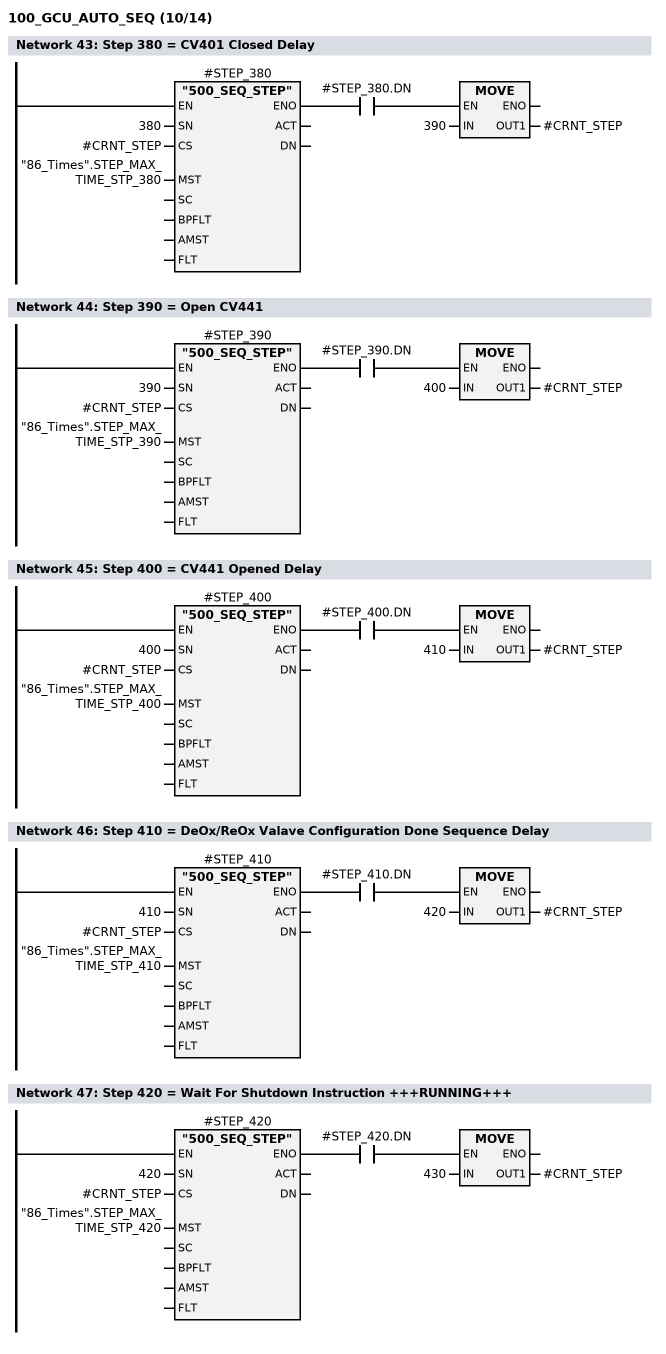
   RUNG wire#powerrail
      #STEP_380(SN := 380, CS := #CRNT_STEP, MST := "86_Times".STEP_MAX_TIME_STP_380, SC :=, BPFLT :=, AMST :=, FLT :=, ACT =>, DN =>)
      Contact( #STEP_380.DN )
      Move(in := 390, out1 => #CRNT_STEP)
   END_RUNG
   // the same network as SCL:
   #STEP_380(SN := 380, CS := #CRNT_STEP, MST := "86_Times".STEP_MAX_TIME_STP_380, ENO => #_w1);   // "500_SEQ_STEP"
   IF #_w1 AND #STEP_380.DN THEN #CRNT_STEP := 390; END_IF;
END_REGION

REGION Network 44: Step 390 = Open CV441
   RUNG wire#powerrail
      #STEP_390(SN := 390, CS := #CRNT_STEP, MST := "86_Times".STEP_MAX_TIME_STP_390, SC :=, BPFLT :=, AMST :=, FLT :=, ACT =>, DN =>)
      Contact( #STEP_390.DN )
      Move(in := 400, out1 => #CRNT_STEP)
   END_RUNG
   // the same network as SCL:
   #STEP_390(SN := 390, CS := #CRNT_STEP, MST := "86_Times".STEP_MAX_TIME_STP_390, ENO => #_w1);   // "500_SEQ_STEP"
   IF #_w1 AND #STEP_390.DN THEN #CRNT_STEP := 400; END_IF;
END_REGION

REGION Network 45: Step 400 = CV441 Opened Delay
   RUNG wire#powerrail
      #STEP_400(SN := 400, CS := #CRNT_STEP, MST := "86_Times".STEP_MAX_TIME_STP_400, SC :=, BPFLT :=, AMST :=, FLT :=, ACT =>, DN =>)
      Contact( #STEP_400.DN )
      Move(in := 410, out1 => #CRNT_STEP)
   END_RUNG
   // the same network as SCL:
   #STEP_400(SN := 400, CS := #CRNT_STEP, MST := "86_Times".STEP_MAX_TIME_STP_400, ENO => #_w1);   // "500_SEQ_STEP"
   IF #_w1 AND #STEP_400.DN THEN #CRNT_STEP := 410; END_IF;
END_REGION

REGION Network 46: Step 410 = DeOx/ReOx Valave Configuration Done Sequence Delay
   RUNG wire#powerrail
      #STEP_410(SN := 410, CS := #CRNT_STEP, MST := "86_Times".STEP_MAX_TIME_STP_410, SC :=, BPFLT :=, AMST :=, FLT :=, ACT =>, DN =>)
      Contact( #STEP_410.DN )
      Move(in := 420, out1 => #CRNT_STEP)
   END_RUNG
   // the same network as SCL:
   #STEP_410(SN := 410, CS := #CRNT_STEP, MST := "86_Times".STEP_MAX_TIME_STP_410, ENO => #_w1);   // "500_SEQ_STEP"
   IF #_w1 AND #STEP_410.DN THEN #CRNT_STEP := 420; END_IF;
END_REGION

REGION Network 47: Step 420 = Wait For Shutdown Instruction +++RUNNING+++
   RUNG wire#powerrail
      #STEP_420(SN := 420, CS := #CRNT_STEP, MST := "86_Times".STEP_MAX_TIME_STP_420, SC :=, BPFLT :=, AMST :=, FLT :=, ACT =>, DN =>)
      Contact( #STEP_420.DN )
      Move(in := 430, out1 => #CRNT_STEP)
   END_RUNG
   // the same network as SCL:
   #STEP_420(SN := 420, CS := #CRNT_STEP, MST := "86_Times".STEP_MAX_TIME_STP_420, ENO => #_w1);   // "500_SEQ_STEP"
   IF #_w1 AND #STEP_420.DN THEN #CRNT_STEP := 430; END_IF;
END_REGION

REGION Network 48: Step 430 = Spare Step (Not Used)
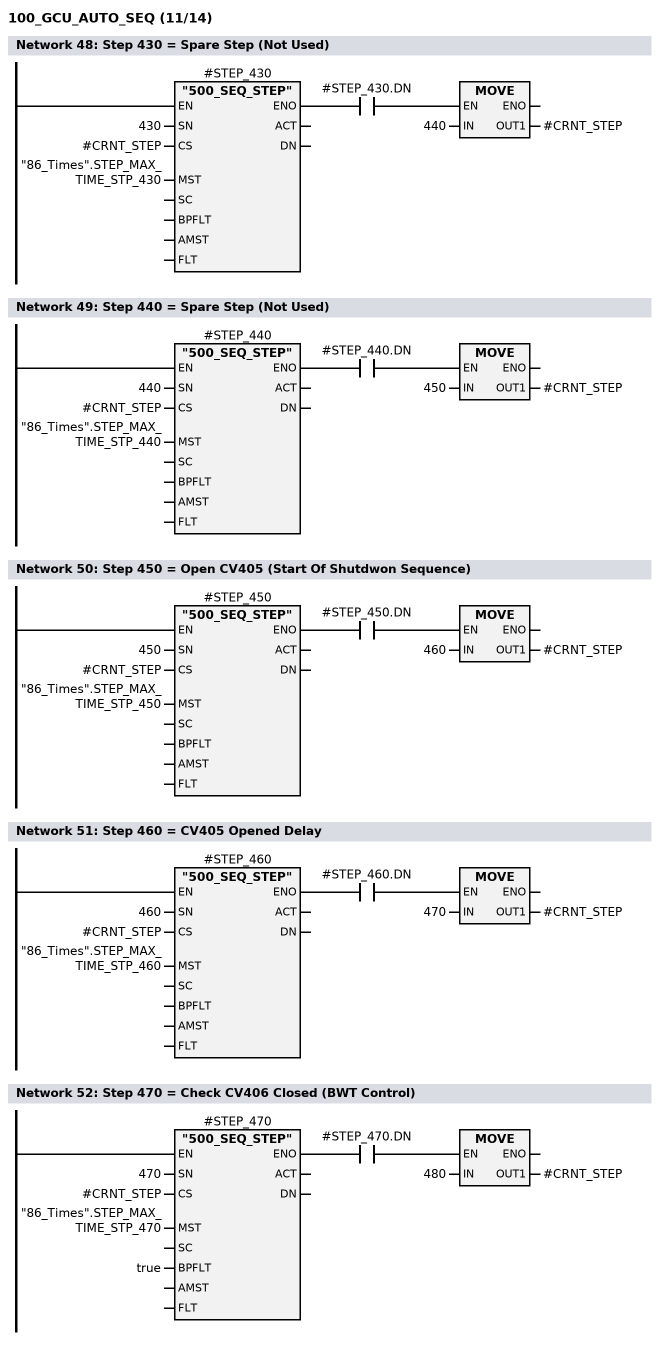
   RUNG wire#powerrail
      #STEP_430(SN := 430, CS := #CRNT_STEP, MST := "86_Times".STEP_MAX_TIME_STP_430, SC :=, BPFLT :=, AMST :=, FLT :=, ACT =>, DN =>)
      Contact( #STEP_430.DN )
      Move(in := 440, out1 => #CRNT_STEP)
   END_RUNG
   // the same network as SCL:
   #STEP_430(SN := 430, CS := #CRNT_STEP, MST := "86_Times".STEP_MAX_TIME_STP_430, ENO => #_w1);   // "500_SEQ_STEP"
   IF #_w1 AND #STEP_430.DN THEN #CRNT_STEP := 440; END_IF;
END_REGION

REGION Network 49: Step 440 = Spare Step (Not Used)
   RUNG wire#powerrail
      #STEP_440(SN := 440, CS := #CRNT_STEP, MST := "86_Times".STEP_MAX_TIME_STP_440, SC :=, BPFLT :=, AMST :=, FLT :=, ACT =>, DN =>)
      Contact( #STEP_440.DN )
      Move(in := 450, out1 => #CRNT_STEP)
   END_RUNG
   // the same network as SCL:
   #STEP_440(SN := 440, CS := #CRNT_STEP, MST := "86_Times".STEP_MAX_TIME_STP_440, ENO => #_w1);   // "500_SEQ_STEP"
   IF #_w1 AND #STEP_440.DN THEN #CRNT_STEP := 450; END_IF;
END_REGION

REGION Network 50: Step 450 = Open CV405 (Start Of Shutdwon Sequence)
   RUNG wire#powerrail
      #STEP_450(SN := 450, CS := #CRNT_STEP, MST := "86_Times".STEP_MAX_TIME_STP_450, SC :=, BPFLT :=, AMST :=, FLT :=, ACT =>, DN =>)
      Contact( #STEP_450.DN )
      Move(in := 460, out1 => #CRNT_STEP)
   END_RUNG
   // the same network as SCL:
   #STEP_450(SN := 450, CS := #CRNT_STEP, MST := "86_Times".STEP_MAX_TIME_STP_450, ENO => #_w1);   // "500_SEQ_STEP"
   IF #_w1 AND #STEP_450.DN THEN #CRNT_STEP := 460; END_IF;
END_REGION

REGION Network 51: Step 460 = CV405 Opened Delay
   RUNG wire#powerrail
      #STEP_460(SN := 460, CS := #CRNT_STEP, MST := "86_Times".STEP_MAX_TIME_STP_460, SC :=, BPFLT :=, AMST :=, FLT :=, ACT =>, DN =>)
      Contact( #STEP_460.DN )
      Move(in := 470, out1 => #CRNT_STEP)
   END_RUNG
   // the same network as SCL:
   #STEP_460(SN := 460, CS := #CRNT_STEP, MST := "86_Times".STEP_MAX_TIME_STP_460, ENO => #_w1);   // "500_SEQ_STEP"
   IF #_w1 AND #STEP_460.DN THEN #CRNT_STEP := 470; END_IF;
END_REGION

REGION Network 52: Step 470 = Check CV406 Closed (BWT Control)
   RUNG wire#powerrail
      #STEP_470(SN := 470, CS := #CRNT_STEP, MST := "86_Times".STEP_MAX_TIME_STP_470, SC :=, BPFLT := true, AMST :=, FLT :=, ACT =>, DN =>)
      Contact( #STEP_470.DN )
      Move(in := 480, out1 => #CRNT_STEP)
   END_RUNG
   // the same network as SCL:
   #STEP_470(SN := 470, CS := #CRNT_STEP, MST := "86_Times".STEP_MAX_TIME_STP_470, BPFLT := true, ENO => #_w1);   // "500_SEQ_STEP"
   IF #_w1 AND #STEP_470.DN THEN #CRNT_STEP := 480; END_IF;
END_REGION

REGION Network 53: Step 480 = CV406 Closed Delay
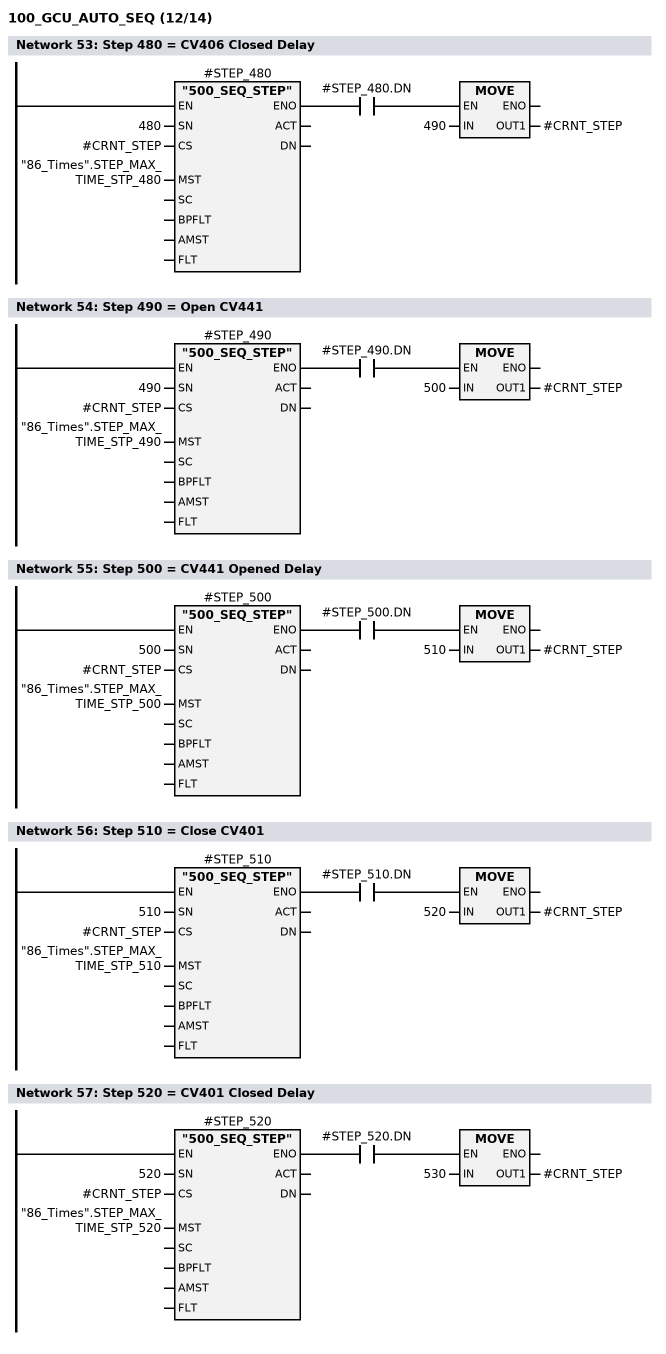
   RUNG wire#powerrail
      #STEP_480(SN := 480, CS := #CRNT_STEP, MST := "86_Times".STEP_MAX_TIME_STP_480, SC :=, BPFLT :=, AMST :=, FLT :=, ACT =>, DN =>)
      Contact( #STEP_480.DN )
      Move(in := 490, out1 => #CRNT_STEP)
   END_RUNG
   // the same network as SCL:
   #STEP_480(SN := 480, CS := #CRNT_STEP, MST := "86_Times".STEP_MAX_TIME_STP_480, ENO => #_w1);   // "500_SEQ_STEP"
   IF #_w1 AND #STEP_480.DN THEN #CRNT_STEP := 490; END_IF;
END_REGION

REGION Network 54: Step 490 = Open CV441
   RUNG wire#powerrail
      #STEP_490(SN := 490, CS := #CRNT_STEP, MST := "86_Times".STEP_MAX_TIME_STP_490, SC :=, BPFLT :=, AMST :=, FLT :=, ACT =>, DN =>)
      Contact( #STEP_490.DN )
      Move(in := 500, out1 => #CRNT_STEP)
   END_RUNG
   // the same network as SCL:
   #STEP_490(SN := 490, CS := #CRNT_STEP, MST := "86_Times".STEP_MAX_TIME_STP_490, ENO => #_w1);   // "500_SEQ_STEP"
   IF #_w1 AND #STEP_490.DN THEN #CRNT_STEP := 500; END_IF;
END_REGION

REGION Network 55: Step 500 = CV441 Opened Delay
   RUNG wire#powerrail
      #STEP_500(SN := 500, CS := #CRNT_STEP, MST := "86_Times".STEP_MAX_TIME_STP_500, SC :=, BPFLT :=, AMST :=, FLT :=, ACT =>, DN =>)
      Contact( #STEP_500.DN )
      Move(in := 510, out1 => #CRNT_STEP)
   END_RUNG
   // the same network as SCL:
   #STEP_500(SN := 500, CS := #CRNT_STEP, MST := "86_Times".STEP_MAX_TIME_STP_500, ENO => #_w1);   // "500_SEQ_STEP"
   IF #_w1 AND #STEP_500.DN THEN #CRNT_STEP := 510; END_IF;
END_REGION

REGION Network 56: Step 510 = Close CV401
   RUNG wire#powerrail
      #STEP_510(SN := 510, CS := #CRNT_STEP, MST := "86_Times".STEP_MAX_TIME_STP_510, SC :=, BPFLT :=, AMST :=, FLT :=, ACT =>, DN =>)
      Contact( #STEP_510.DN )
      Move(in := 520, out1 => #CRNT_STEP)
   END_RUNG
   // the same network as SCL:
   #STEP_510(SN := 510, CS := #CRNT_STEP, MST := "86_Times".STEP_MAX_TIME_STP_510, ENO => #_w1);   // "500_SEQ_STEP"
   IF #_w1 AND #STEP_510.DN THEN #CRNT_STEP := 520; END_IF;
END_REGION

REGION Network 57: Step 520 = CV401 Closed Delay
   RUNG wire#powerrail
      #STEP_520(SN := 520, CS := #CRNT_STEP, MST := "86_Times".STEP_MAX_TIME_STP_520, SC :=, BPFLT :=, AMST :=, FLT :=, ACT =>, DN =>)
      Contact( #STEP_520.DN )
      Move(in := 530, out1 => #CRNT_STEP)
   END_RUNG
   // the same network as SCL:
   #STEP_520(SN := 520, CS := #CRNT_STEP, MST := "86_Times".STEP_MAX_TIME_STP_520, ENO => #_w1);   // "500_SEQ_STEP"
   IF #_w1 AND #STEP_520.DN THEN #CRNT_STEP := 530; END_IF;
END_REGION

REGION Network 58: Step 530 = Stop E400
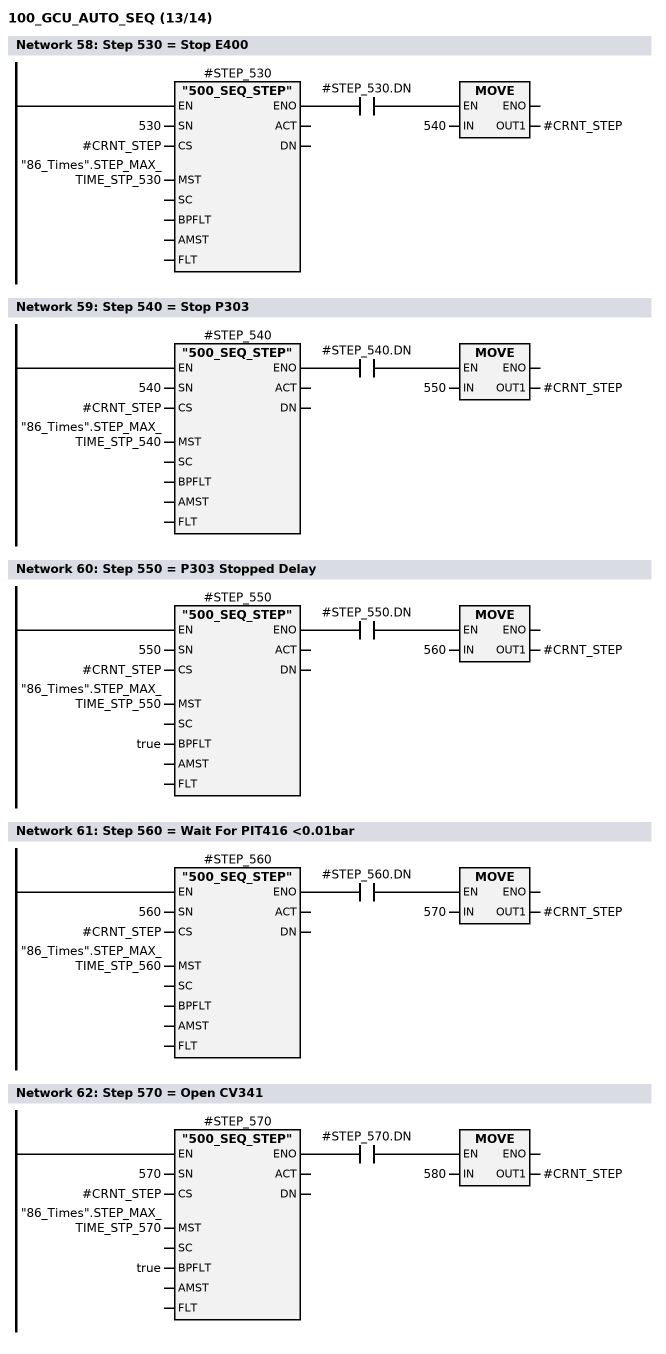
   RUNG wire#powerrail
      #STEP_530(SN := 530, CS := #CRNT_STEP, MST := "86_Times".STEP_MAX_TIME_STP_530, SC :=, BPFLT :=, AMST :=, FLT :=, ACT =>, DN =>)
      Contact( #STEP_530.DN )
      Move(in := 540, out1 => #CRNT_STEP)
   END_RUNG
   // the same network as SCL:
   #STEP_530(SN := 530, CS := #CRNT_STEP, MST := "86_Times".STEP_MAX_TIME_STP_530, ENO => #_w1);   // "500_SEQ_STEP"
   IF #_w1 AND #STEP_530.DN THEN #CRNT_STEP := 540; END_IF;
END_REGION

REGION Network 59: Step 540 = Stop P303
   RUNG wire#powerrail
      #STEP_540(SN := 540, CS := #CRNT_STEP, MST := "86_Times".STEP_MAX_TIME_STP_540, SC :=, BPFLT :=, AMST :=, FLT :=, ACT =>, DN =>)
      Contact( #STEP_540.DN )
      Move(in := 550, out1 => #CRNT_STEP)
   END_RUNG
   // the same network as SCL:
   #STEP_540(SN := 540, CS := #CRNT_STEP, MST := "86_Times".STEP_MAX_TIME_STP_540, ENO => #_w1);   // "500_SEQ_STEP"
   IF #_w1 AND #STEP_540.DN THEN #CRNT_STEP := 550; END_IF;
END_REGION

REGION Network 60: Step 550 = P303 Stopped Delay
   RUNG wire#powerrail
      #STEP_550(SN := 550, CS := #CRNT_STEP, MST := "86_Times".STEP_MAX_TIME_STP_550, SC :=, BPFLT := true, AMST :=, FLT :=, ACT =>, DN =>)
      Contact( #STEP_550.DN )
      Move(in := 560, out1 => #CRNT_STEP)
   END_RUNG
   // the same network as SCL:
   #STEP_550(SN := 550, CS := #CRNT_STEP, MST := "86_Times".STEP_MAX_TIME_STP_550, BPFLT := true, ENO => #_w1);   // "500_SEQ_STEP"
   IF #_w1 AND #STEP_550.DN THEN #CRNT_STEP := 560; END_IF;
END_REGION

REGION Network 61: Step 560 = Wait For PIT416 <0.01bar
   RUNG wire#powerrail
      #STEP_560(SN := 560, CS := #CRNT_STEP, MST := "86_Times".STEP_MAX_TIME_STP_560, SC :=, BPFLT :=, AMST :=, FLT :=, ACT =>, DN =>)
      Contact( #STEP_560.DN )
      Move(in := 570, out1 => #CRNT_STEP)
   END_RUNG
   // the same network as SCL:
   #STEP_560(SN := 560, CS := #CRNT_STEP, MST := "86_Times".STEP_MAX_TIME_STP_560, ENO => #_w1);   // "500_SEQ_STEP"
   IF #_w1 AND #STEP_560.DN THEN #CRNT_STEP := 570; END_IF;
END_REGION

REGION Network 62: Step 570 = Open CV341
   RUNG wire#powerrail
      #STEP_570(SN := 570, CS := #CRNT_STEP, MST := "86_Times".STEP_MAX_TIME_STP_570, SC :=, BPFLT := true, AMST :=, FLT :=, ACT =>, DN =>)
      Contact( #STEP_570.DN )
      Move(in := 580, out1 => #CRNT_STEP)
   END_RUNG
   // the same network as SCL:
   #STEP_570(SN := 570, CS := #CRNT_STEP, MST := "86_Times".STEP_MAX_TIME_STP_570, BPFLT := true, ENO => #_w1);   // "500_SEQ_STEP"
   IF #_w1 AND #STEP_570.DN THEN #CRNT_STEP := 580; END_IF;
END_REGION

REGION Network 63: Step 580 = CV341 Opened Delay
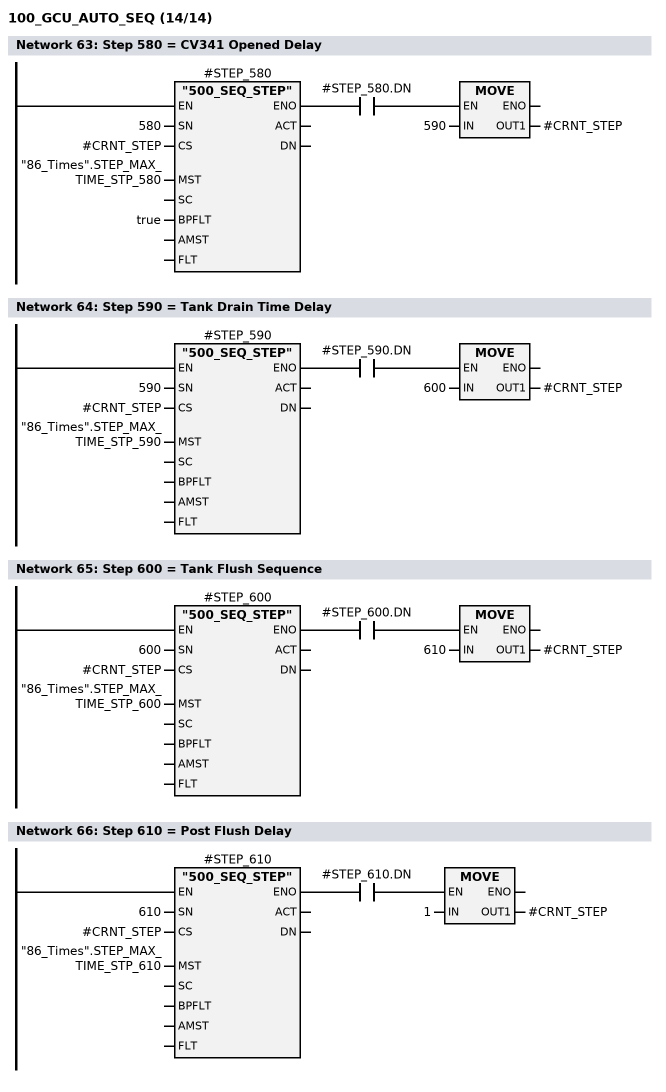
   RUNG wire#powerrail
      #STEP_580(SN := 580, CS := #CRNT_STEP, MST := "86_Times".STEP_MAX_TIME_STP_580, SC :=, BPFLT := true, AMST :=, FLT :=, ACT =>, DN =>)
      Contact( #STEP_580.DN )
      Move(in := 590, out1 => #CRNT_STEP)
   END_RUNG
   // the same network as SCL:
   #STEP_580(SN := 580, CS := #CRNT_STEP, MST := "86_Times".STEP_MAX_TIME_STP_580, BPFLT := true, ENO => #_w1);   // "500_SEQ_STEP"
   IF #_w1 AND #STEP_580.DN THEN #CRNT_STEP := 590; END_IF;
END_REGION

REGION Network 64: Step 590 = Tank Drain Time Delay
   RUNG wire#powerrail
      #STEP_590(SN := 590, CS := #CRNT_STEP, MST := "86_Times".STEP_MAX_TIME_STP_590, SC :=, BPFLT :=, AMST :=, FLT :=, ACT =>, DN =>)
      Contact( #STEP_590.DN )
      Move(in := 600, out1 => #CRNT_STEP)
   END_RUNG
   // the same network as SCL:
   #STEP_590(SN := 590, CS := #CRNT_STEP, MST := "86_Times".STEP_MAX_TIME_STP_590, ENO => #_w1);   // "500_SEQ_STEP"
   IF #_w1 AND #STEP_590.DN THEN #CRNT_STEP := 600; END_IF;
END_REGION

REGION Network 65: Step 600 = Tank Flush Sequence
   RUNG wire#powerrail
      #STEP_600(SN := 600, CS := #CRNT_STEP, MST := "86_Times".STEP_MAX_TIME_STP_600, SC :=, BPFLT :=, AMST :=, FLT :=, ACT =>, DN =>)
      Contact( #STEP_600.DN )
      Move(in := 610, out1 => #CRNT_STEP)
   END_RUNG
   // the same network as SCL:
   #STEP_600(SN := 600, CS := #CRNT_STEP, MST := "86_Times".STEP_MAX_TIME_STP_600, ENO => #_w1);   // "500_SEQ_STEP"
   IF #_w1 AND #STEP_600.DN THEN #CRNT_STEP := 610; END_IF;
END_REGION

REGION Network 66: Step 610 = Post Flush Delay
   RUNG wire#powerrail
      #STEP_610(SN := 610, CS := #CRNT_STEP, MST := "86_Times".STEP_MAX_TIME_STP_610, SC :=, BPFLT :=, AMST :=, FLT :=, ACT =>, DN =>)
      Contact( #STEP_610.DN )
      Move(in := 1, out1 => #CRNT_STEP)
   END_RUNG
   // the same network as SCL:
   #STEP_610(SN := 610, CS := #CRNT_STEP, MST := "86_Times".STEP_MAX_TIME_STP_610, ENO => #_w1);   // "500_SEQ_STEP"
   IF #_w1 AND #STEP_610.DN THEN #CRNT_STEP := 1; END_IF;
END_REGION
END_FUNCTION_BLOCK

FUNCTION_BLOCK "Setpoint Override"   // FB104, LAD
{ S7_Optimized_Access := 'TRUE' }
VERSION : 0.1
   VAR_INPUT
      Enable : Bool;
      "Activate Temp Prot" : Bool := true;
      Temperature : Real;
      "Temperature Setpoint" : Real := 250.0;
      "Temperature Tolerance" : Real := 10.0;
      "Activate Press Prot" : Bool;
      Pressure : Real;
      "Pressure Setpoint" : Real := 5.0;
      "Pressure Tolerance" : Real := 0.2;
      "Pressure Target" : Real := 3.5;
      "Pressure Safe Target" : Real := 3.0;
      "Activate Tank Change Prot" : Bool := true;
      "Tank Change TimeOut" : Time := T#60s;
      "Tank Change" : Bool := true;
      Reset : Bool;
   END_VAR
   VAR_OUTPUT
      "Pressure Target Override" : Real;
      "Pressure Safe Override" : Real;
   END_VAR
   VAR
      "Temperature Setpoint Aux" : Real;
      "Pressure Setpoint Aux" : Real;
      "Set Pressure" : Bool;
      "Set Pressure Aux" : Bool;
      "Set Pressure by Temp" : Bool;
      "Set Pressure by Press" : Bool;
      "Set Pressure by Tank" : Bool;
   END_VAR
   VAR RETAIN
      "Pressure Target Memory" : Real;
   END_VAR
   VAR
      "Set Pressure Puls1" : Bool;
      "Set Pressure Puls2" : Bool;
      "Tank Change Protection" : TOF_TIME;
      "Pressure Protection" : TOF_TIME;
      "Pressure Memory Recover" : TON_TIME;
   END_VAR
   VAR_TEMP   // added for the SCL form of the ladder/FBD networks
      _w1 : Bool;
   END_VAR
BEGIN

REGION Network 1: Pressure Safe Corection
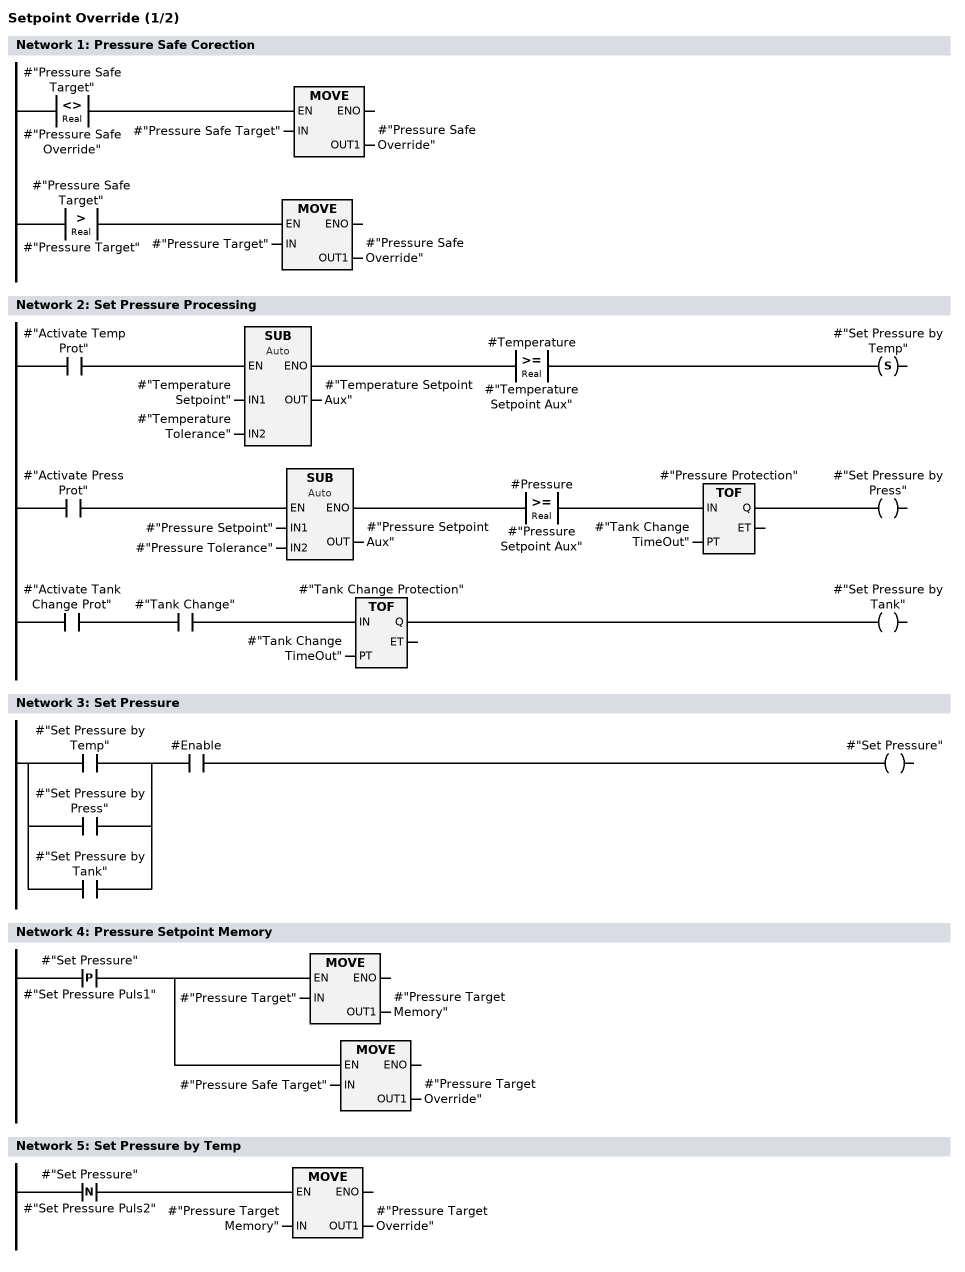
   RUNG wire#powerrail
      { S7_Templates := "SrcType := Real" } NE_Contact(in1 := #"Pressure Safe Target", in2 := #"Pressure Safe Override")
      Move(in := #"Pressure Safe Target", out1 => #"Pressure Safe Override")
   END_RUNG
   RUNG wire#powerrail
      { S7_Templates := "SrcType := Real" } GT_Contact(in1 := #"Pressure Safe Target", in2 := #"Pressure Target")
      Move(in := #"Pressure Target", out1 => #"Pressure Safe Override")
   END_RUNG
   // the same network as SCL:
   IF #"Pressure Safe Target" <> #"Pressure Safe Override" THEN
       #"Pressure Safe Override" := #"Pressure Safe Target";
   END_IF;
   IF #"Pressure Safe Target" > #"Pressure Target" THEN
       #"Pressure Safe Override" := #"Pressure Target";
   END_IF;
END_REGION

REGION Network 2: Set Pressure Processing
   IF #"Activate Temp Prot" THEN
       #"Temperature Setpoint Aux" := #"Temperature Setpoint" - #"Temperature Tolerance";
   END_IF;
   IF #"Activate Temp Prot" AND (#Temperature >= #"Temperature Setpoint Aux") THEN
       #"Set Pressure by Temp" := TRUE;
   END_IF;
   IF #"Activate Press Prot" THEN
       #"Pressure Setpoint Aux" := #"Pressure Setpoint" - #"Pressure Tolerance";
   END_IF;
   #"Pressure Protection"(IN := #"Activate Press Prot" AND (#Pressure >= #"Pressure Setpoint Aux"),   // TOF
                          PT := #"Tank Change TimeOut");
   #"Set Pressure by Press" := #"Pressure Protection".Q;
   #"Tank Change Protection"(IN := #"Activate Tank Change Prot" AND #"Tank Change",   // TOF
                           PT := #"Tank Change TimeOut");
   #"Set Pressure by Tank" := #"Tank Change Protection".Q;
END_REGION

REGION Network 3: Set Pressure
   RUNG wire#powerrail
      Contact( #"Set Pressure by Temp" )
      wire#w1
      Contact( #Enable )
      Coil( #"Set Pressure" )
   END_RUNG
   RUNG wire#powerrail
      Contact( #"Set Pressure by Press" )
   END_RUNG wire#w1
   RUNG wire#powerrail
      Contact( #"Set Pressure by Tank" )
   END_RUNG wire#w1
   // the same network as SCL:
   #"Set Pressure" := (#"Set Pressure by Temp" OR #"Set Pressure by Press" OR #"Set Pressure by Tank") AND #Enable;
END_REGION

REGION Network 4: Pressure Setpoint Memory
   RUNG wire#powerrail
      P_Contact(operand := #"Set Pressure", bit := #"Set Pressure Puls1")
      wire#w1
      Move(in := #"Pressure Target", out1 => #"Pressure Target Memory")
   END_RUNG
   RUNG wire#w1
      Move(in := #"Pressure Safe Target", out1 => #"Pressure Target Override")
   END_RUNG
   // the same network as SCL:
   #_w1 := #"Set Pressure" AND NOT #"Set Pressure Puls1";   // rising edge of #"Set Pressure"
   #"Set Pressure Puls1" := #"Set Pressure";
   IF #_w1 THEN
       #"Pressure Target Memory" := #"Pressure Target";
       #"Pressure Target Override" := #"Pressure Safe Target";
   END_IF;
END_REGION

REGION Network 5: Set Pressure by Temp
   RUNG wire#powerrail
      N_Contact(operand := #"Set Pressure", bit := #"Set Pressure Puls2")
      Move(in := #"Pressure Target Memory", out1 => #"Pressure Target Override")
   END_RUNG
   // the same network as SCL:
   #_w1 := NOT #"Set Pressure" AND #"Set Pressure Puls2";   // falling edge of #"Set Pressure"
   #"Set Pressure Puls2" := #"Set Pressure";
   IF #_w1 THEN #"Pressure Target Override" := #"Pressure Target Memory"; END_IF;
END_REGION

REGION Network 6: Set Pressure Back
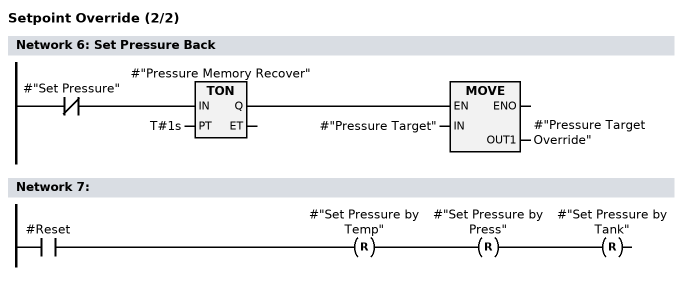
   #"Pressure Memory Recover"(IN := NOT #"Set Pressure", PT := T#1s);   // TON
   IF #"Pressure Memory Recover".Q THEN #"Pressure Target Override" := #"Pressure Target"; END_IF;
END_REGION

REGION Network 7
   RUNG wire#powerrail
      Contact( #Reset )
      R_Coil( #"Set Pressure by Temp" )
      R_Coil( #"Set Pressure by Press" )
      R_Coil( #"Set Pressure by Tank" )
   END_RUNG
   // the same network as SCL:
   IF #Reset THEN
       #"Set Pressure by Temp" := FALSE;
       #"Set Pressure by Press" := FALSE;
       #"Set Pressure by Tank" := FALSE;
   END_IF;
END_REGION
END_FUNCTION_BLOCK

FUNCTION_BLOCK "108_GCU_TNK_REFILL_SEQ"   // FB108, LAD
TITLE = GCU Tank Refill Sequence
{ S7_Optimized_Access := 'TRUE' }
AUTHOR : JRS
VERSION : 0.1
// For the automatic refilling of the GCU tank to the required level
   VAR_INPUT
      RUN : Bool;   // Block control
      LEVEL : Real;   // Tank level value
      TARGET : Real;   // Target level value
      LOW : Real;   // Low level value
      P305_PRSNT : Bool;   // P305 Fitted
      P305_RNG : Bool;   // Pump running
      P304_RNG : Bool;   // Pump running
      CV358_OPN : Bool;   // Valve open
      CV358_CLSD : Bool;   // Valve closed
   END_VAR
   VAR_OUTPUT
      RUN_P305 : Bool;   // Pump control
      RUN_P304 : Bool;   // Pump control
      OPEN_CV358 : Bool;   // Valve control
      FILLING : Bool;   // Filling status
   END_VAR
   VAR
      INTO_RUN_PLS : Bool;   // Pulse bit
      "STEP" : Int;   // Step number
      RNG : Bool;   // Running bit
      OUT_RUN_PLS : Bool;   // Pulse bit
   END_VAR
   VAR_TEMP   // added for the SCL form of the ladder/FBD networks
      _w1 : Bool;
   END_VAR
BEGIN

REGION Network 1: First Into Run
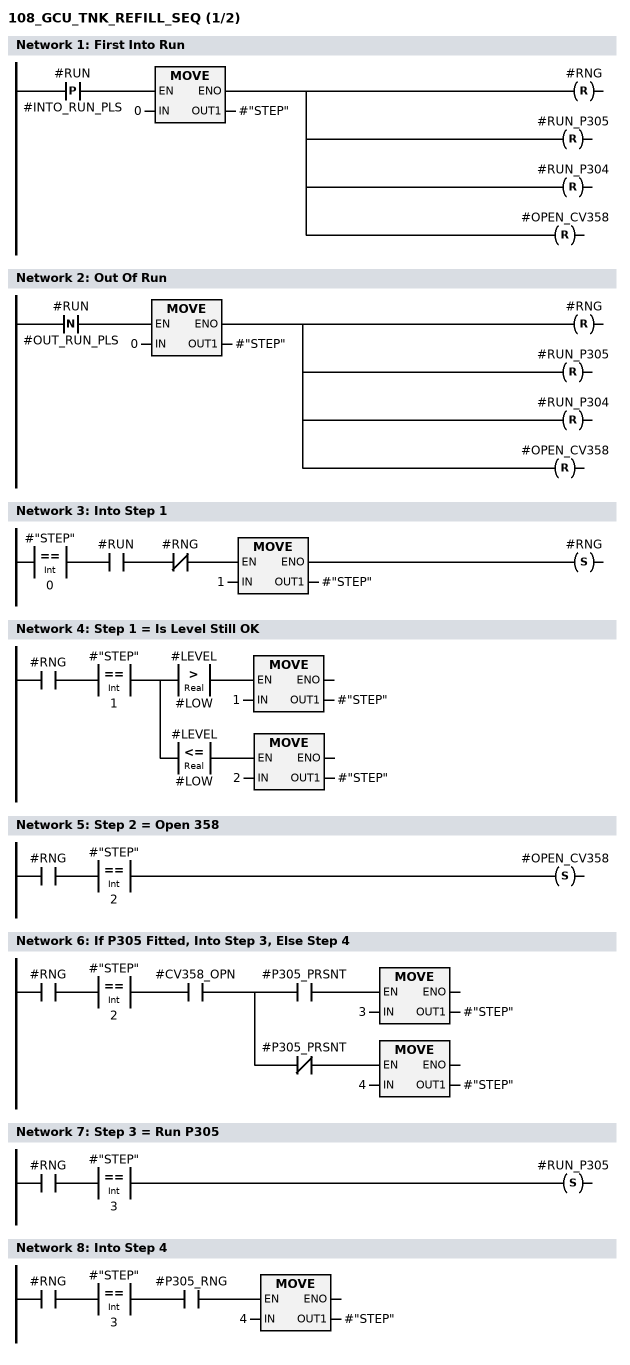
   RUNG wire#powerrail
      P_Contact(operand := #RUN, bit := #INTO_RUN_PLS)
      Move(in := 0, out1 => #"STEP")
      wire#w1
      R_Coil( #RNG )
   END_RUNG
   RUNG wire#w1
      R_Coil( #RUN_P305 )
   END_RUNG
   RUNG wire#w1
      R_Coil( #RUN_P304 )
   END_RUNG
   RUNG wire#w1
      R_Coil( #OPEN_CV358 )
   END_RUNG
   // the same network as SCL:
   #_w1 := #RUN AND NOT #INTO_RUN_PLS;   // rising edge of #RUN
   #INTO_RUN_PLS := #RUN;
   IF #_w1 THEN
       #"STEP" := 0;
       #RNG := FALSE;
       #RUN_P305 := FALSE;
       #RUN_P304 := FALSE;
       #OPEN_CV358 := FALSE;
   END_IF;
END_REGION

REGION Network 2: Out Of Run
   RUNG wire#powerrail
      N_Contact(operand := #RUN, bit := #OUT_RUN_PLS)
      Move(in := 0, out1 => #"STEP")
      wire#w1
      R_Coil( #RNG )
   END_RUNG
   RUNG wire#w1
      R_Coil( #RUN_P305 )
   END_RUNG
   RUNG wire#w1
      R_Coil( #RUN_P304 )
   END_RUNG
   RUNG wire#w1
      R_Coil( #OPEN_CV358 )
   END_RUNG
   // the same network as SCL:
   #_w1 := NOT #RUN AND #OUT_RUN_PLS;   // falling edge of #RUN
   #OUT_RUN_PLS := #RUN;
   IF #_w1 THEN
       #"STEP" := 0;
       #RNG := FALSE;
       #RUN_P305 := FALSE;
       #RUN_P304 := FALSE;
       #OPEN_CV358 := FALSE;
   END_IF;
END_REGION

REGION Network 3: Into Step 1
   RUNG wire#powerrail
      { S7_Templates := "SrcType := Int" } EQ_Contact(in1 := #"STEP", in2 := 0)
      Contact( #RUN )
      I_Contact( #RNG )
      Move(in := 1, out1 => #"STEP")
      S_Coil( #RNG )
   END_RUNG
   // the same network as SCL:
   #_w1 := (#"STEP" = 0) AND #RUN AND NOT #RNG;
   IF #_w1 THEN
       #"STEP" := 1;
       #RNG := TRUE;
   END_IF;
END_REGION

REGION Network 4: Step 1 = Is Level Still OK
   RUNG wire#powerrail
      Contact( #RNG )
      { S7_Templates := "SrcType := Int" } EQ_Contact(in1 := #"STEP", in2 := 1)
      wire#w1
      { S7_Templates := "SrcType := Real" } GT_Contact(in1 := #LEVEL, in2 := #LOW)
      Move(in := 1, out1 => #"STEP")
   END_RUNG
   RUNG wire#w1
      { S7_Templates := "SrcType := Real" } LE_Contact(in1 := #LEVEL, in2 := #LOW)
      Move(in := 2, out1 => #"STEP")
   END_RUNG
   // the same network as SCL:
   #_w1 := #RNG AND (#"STEP" = 1);
   IF #_w1 AND (#LEVEL > #LOW) THEN #"STEP" := 1; END_IF;
   IF #_w1 AND (#LEVEL <= #LOW) THEN #"STEP" := 2; END_IF;
END_REGION

REGION Network 5: Step 2 = Open 358
   RUNG wire#powerrail
      Contact( #RNG )
      { S7_Templates := "SrcType := Int" } EQ_Contact(in1 := #"STEP", in2 := 2)
      S_Coil( #OPEN_CV358 )
   END_RUNG
   // the same network as SCL:
   IF #RNG AND (#"STEP" = 2) THEN #OPEN_CV358 := TRUE; END_IF;
END_REGION

REGION Network 6: If P305 Fitted, Into Step 3, Else Step 4
   RUNG wire#powerrail
      Contact( #RNG )
      { S7_Templates := "SrcType := Int" } EQ_Contact(in1 := #"STEP", in2 := 2)
      Contact( #CV358_OPN )
      wire#w1
      Contact( #P305_PRSNT )
      Move(in := 3, out1 => #"STEP")
   END_RUNG
   RUNG wire#w1
      I_Contact( #P305_PRSNT )
      Move(in := 4, out1 => #"STEP")
   END_RUNG
   // the same network as SCL:
   #_w1 := #RNG AND (#"STEP" = 2) AND #CV358_OPN;
   IF #_w1 AND #P305_PRSNT THEN #"STEP" := 3; END_IF;
   IF #_w1 AND NOT #P305_PRSNT THEN #"STEP" := 4; END_IF;
END_REGION

REGION Network 7: Step 3 = Run P305
   RUNG wire#powerrail
      Contact( #RNG )
      { S7_Templates := "SrcType := Int" } EQ_Contact(in1 := #"STEP", in2 := 3)
      S_Coil( #RUN_P305 )
   END_RUNG
   // the same network as SCL:
   IF #RNG AND (#"STEP" = 3) THEN #RUN_P305 := TRUE; END_IF;
END_REGION

REGION Network 8: Into Step 4
   RUNG wire#powerrail
      Contact( #RNG )
      { S7_Templates := "SrcType := Int" } EQ_Contact(in1 := #"STEP", in2 := 3)
      Contact( #P305_RNG )
      Move(in := 4, out1 => #"STEP")
   END_RUNG
   // the same network as SCL:
   IF #RNG AND (#"STEP" = 3) AND #P305_RNG THEN #"STEP" := 4; END_IF;
END_REGION

REGION Network 9: Step 4 = Run P304
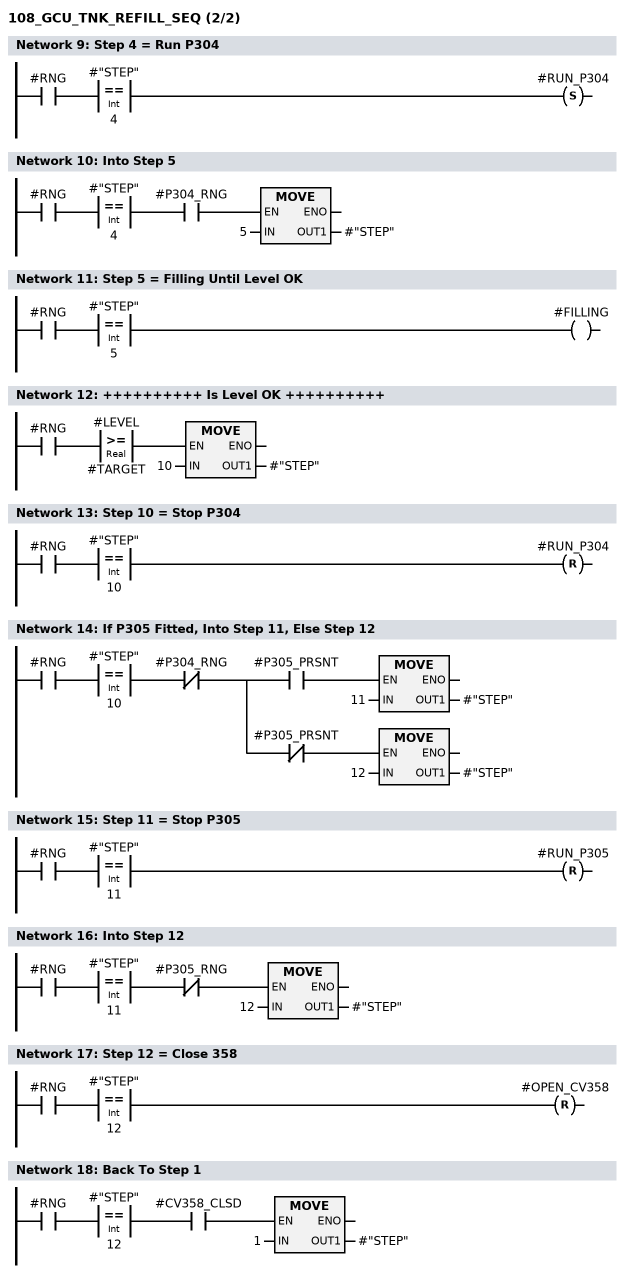
   RUNG wire#powerrail
      Contact( #RNG )
      { S7_Templates := "SrcType := Int" } EQ_Contact(in1 := #"STEP", in2 := 4)
      S_Coil( #RUN_P304 )
   END_RUNG
   // the same network as SCL:
   IF #RNG AND (#"STEP" = 4) THEN #RUN_P304 := TRUE; END_IF;
END_REGION

REGION Network 10: Into Step 5
   RUNG wire#powerrail
      Contact( #RNG )
      { S7_Templates := "SrcType := Int" } EQ_Contact(in1 := #"STEP", in2 := 4)
      Contact( #P304_RNG )
      Move(in := 5, out1 => #"STEP")
   END_RUNG
   // the same network as SCL:
   IF #RNG AND (#"STEP" = 4) AND #P304_RNG THEN #"STEP" := 5; END_IF;
END_REGION

REGION Network 11: Step 5 = Filling Until Level OK
   RUNG wire#powerrail
      Contact( #RNG )
      { S7_Templates := "SrcType := Int" } EQ_Contact(in1 := #"STEP", in2 := 5)
      Coil( #FILLING )
   END_RUNG
   // the same network as SCL:
   #FILLING := #RNG AND (#"STEP" = 5);
END_REGION

REGION Network 12: ++++++++++ Is Level OK ++++++++++
   RUNG wire#powerrail
      Contact( #RNG )
      { S7_Templates := "SrcType := Real" } GE_Contact(in1 := #LEVEL, in2 := #TARGET)
      Move(in := 10, out1 => #"STEP")
   END_RUNG
   // the same network as SCL:
   IF #RNG AND (#LEVEL >= #TARGET) THEN #"STEP" := 10; END_IF;
END_REGION

REGION Network 13: Step 10 = Stop P304
   RUNG wire#powerrail
      Contact( #RNG )
      { S7_Templates := "SrcType := Int" } EQ_Contact(in1 := #"STEP", in2 := 10)
      R_Coil( #RUN_P304 )
   END_RUNG
   // the same network as SCL:
   IF #RNG AND (#"STEP" = 10) THEN #RUN_P304 := FALSE; END_IF;
END_REGION

REGION Network 14: If P305 Fitted, Into Step 11, Else Step 12
   RUNG wire#powerrail
      Contact( #RNG )
      { S7_Templates := "SrcType := Int" } EQ_Contact(in1 := #"STEP", in2 := 10)
      I_Contact( #P304_RNG )
      wire#w1
      Contact( #P305_PRSNT )
      Move(in := 11, out1 => #"STEP")
   END_RUNG
   RUNG wire#w1
      I_Contact( #P305_PRSNT )
      Move(in := 12, out1 => #"STEP")
   END_RUNG
   // the same network as SCL:
   #_w1 := #RNG AND (#"STEP" = 10) AND NOT #P304_RNG;
   IF #_w1 AND #P305_PRSNT THEN #"STEP" := 11; END_IF;
   IF #_w1 AND NOT #P305_PRSNT THEN #"STEP" := 12; END_IF;
END_REGION

REGION Network 15: Step 11 = Stop P305
   RUNG wire#powerrail
      Contact( #RNG )
      { S7_Templates := "SrcType := Int" } EQ_Contact(in1 := #"STEP", in2 := 11)
      R_Coil( #RUN_P305 )
   END_RUNG
   // the same network as SCL:
   IF #RNG AND (#"STEP" = 11) THEN #RUN_P305 := FALSE; END_IF;
END_REGION

REGION Network 16: Into Step 12
   RUNG wire#powerrail
      Contact( #RNG )
      { S7_Templates := "SrcType := Int" } EQ_Contact(in1 := #"STEP", in2 := 11)
      I_Contact( #P305_RNG )
      Move(in := 12, out1 => #"STEP")
   END_RUNG
   // the same network as SCL:
   IF #RNG AND (#"STEP" = 11) AND NOT #P305_RNG THEN #"STEP" := 12; END_IF;
END_REGION

REGION Network 17: Step 12 = Close 358
   RUNG wire#powerrail
      Contact( #RNG )
      { S7_Templates := "SrcType := Int" } EQ_Contact(in1 := #"STEP", in2 := 12)
      R_Coil( #OPEN_CV358 )
   END_RUNG
   // the same network as SCL:
   IF #RNG AND (#"STEP" = 12) THEN #OPEN_CV358 := FALSE; END_IF;
END_REGION

REGION Network 18: Back To Step 1
   RUNG wire#powerrail
      Contact( #RNG )
      { S7_Templates := "SrcType := Int" } EQ_Contact(in1 := #"STEP", in2 := 12)
      Contact( #CV358_CLSD )
      Move(in := 1, out1 => #"STEP")
   END_RUNG
   // the same network as SCL:
   IF #RNG AND (#"STEP" = 12) AND #CV358_CLSD THEN #"STEP" := 1; END_IF;
END_REGION
END_FUNCTION_BLOCK

FUNCTION_BLOCK "109_TRGT_RAMP_CNTRL"   // FB109, LAD
TITLE = Target Control Ramp
{ S7_Optimized_Access := 'TRUE' }
AUTHOR : JRS
VERSION : 0.1
// For the control of target setpoint ramp over specified time
   VAR_INPUT
      RUN : Bool;   // Runs the block
      PRSR : Real;   // Measured preasure level
      TRGT : Real;   // End target value
      "TIME" : Real;   // Ramp time in seconds
   END_VAR
   VAR_OUTPUT
      CMND_TRGT : Real;   // Target value to PID
      DONE : Bool;   // Ramp Done
   END_VAR
   VAR
      "Step" : Int;   // State value for sequencing
      INTO_RUN_PLS : Bool;   // Edge detection
      OUT_RUN_PLS : Bool;   // Edge detection
      RNG : Bool;   // Running
      INIT_PRESS : Real;   // Initial Pressure Level
      DEV_PER_SEC : Real;   // Deveation per second
      UPR_TOL : Real;   // Target + Dev Per Sec
      LWR_TOL : Real;   // Target - Dev Per Sec
      CLK_UP_PLS : Bool;   // Pulse bit
      CLK_DN_PLS : Bool;   // Pulse bit
      CRNT_TRGT : Real;   // Current target
   END_VAR
   VAR_TEMP   // added for the SCL form of the ladder/FBD networks
      _w1 : Bool;
   END_VAR
BEGIN

REGION Network 1: First Into Run